FUNCTION_BLOCK "FB_GL_PROGRAM"   // FB5, GRAPH_PLUS
{ S7_Optimized_Access := 'TRUE' }
VERSION : 0.1
   VAR_INPUT
      OFF_SQ : Bool := false;   // Turn sequence off
      INIT_SQ : Bool := false;   // Set sequence to initial state
      ACK_EF : Bool := false;   // Acknowledge all errors and faults
      S_PREV : Bool := false;   // Output previous step in parameter S_NO
      S_NEXT : Bool := false;   // Indicate next step in parameter S_NO
      SW_AUTO : Bool := false;   // Automatic mode
      SW_TAP : Bool := false;   // Semiautomatic/switch with transition
      SW_TOP : Bool := false;   // Semiautomatic/ignore transition
      SW_MAN : Bool := false;   // Manual mode
      S_SEL : Int := 0;   // Select step to be output to S_NO
      S_ON : Bool := false;   // Activate step indicated in S_NO
      S_OFF : Bool := false;   // Deactivate step indicated S_NO
      T_PUSH : Bool := false;   // Enable transition to switch in semi automatic mode
   END_VAR
   VAR_OUTPUT
      S_NO : Int := 0;   // Step number
      S_MORE : Bool := false;   // More steps are available and can be shown in S_NO
      S_ACTIVE : Bool := false;   // Step indicated in S_NO is active
      ERR_FLT : Bool := false;   // Interlock or supervision group error
      AUTO_ON : Bool := false;   // Automatic mode is active
      TAP_ON : Bool := false;   // Semiautomatic mode/step with transition enabled
      TOP_ON : Bool := false;   // Semiautomatic mode/ignore transition enabled
      MAN_ON : Bool := false;   // Manual mode is active
   END_VAR
   VAR
      T_ON : Array[0..125] of TON_TIME;
   END_VAR
   VAR RETAIN
      StevecKosov : DInt;
   END_VAR
   VAR
      HMI_INFO : Array[0..34] of UInt;
      IF_PAR : G7_IfParPlus_V6;
      RT_DATA : G7_RTDataPlus_V6;   // Internal data area
      Trans9 : G7_TransitionPlus_V6;   // Transition structure
      Trans18 : G7_TransitionPlus_V6;   // Transition structure
      Trans19 : G7_TransitionPlus_V6;   // Transition structure
      Trans20 : G7_TransitionPlus_V6;   // Transition structure
      Trans22 : G7_TransitionPlus_V6;   // Transition structure
      Trans23 : G7_TransitionPlus_V6;   // Transition structure
      Trans24 : G7_TransitionPlus_V6;   // Transition structure
      Trans26 : G7_TransitionPlus_V6;   // Transition structure
      Trans28 : G7_TransitionPlus_V6;   // Transition structure
      Trans29 : G7_TransitionPlus_V6;   // Transition structure
      Trans30 : G7_TransitionPlus_V6;   // Transition structure
      Trans31 : G7_TransitionPlus_V6;   // Transition structure
      Trans32 : G7_TransitionPlus_V6;   // Transition structure
      Trans33 : G7_TransitionPlus_V6;   // Transition structure
      Trans34 : G7_TransitionPlus_V6;   // Transition structure
      Trans35 : G7_TransitionPlus_V6;   // Transition structure
      Trans36 : G7_TransitionPlus_V6;   // Transition structure
      Trans37 : G7_TransitionPlus_V6;   // Transition structure
      Trans38 : G7_TransitionPlus_V6;   // Transition structure
      Trans39 : G7_TransitionPlus_V6;   // Transition structure
      Trans40 : G7_TransitionPlus_V6;   // Transition structure
      Trans41 : G7_TransitionPlus_V6;   // Transition structure
      Trans42 : G7_TransitionPlus_V6;   // Transition structure
      Trans43 : G7_TransitionPlus_V6;   // Transition structure
      Trans44 : G7_TransitionPlus_V6;   // Transition structure
      Trans45 : G7_TransitionPlus_V6;   // Transition structure
      Trans46 : G7_TransitionPlus_V6;   // Transition structure
      Trans47 : G7_TransitionPlus_V6;   // Transition structure
      Trans48 : G7_TransitionPlus_V6;   // Transition structure
      Trans49 : G7_TransitionPlus_V6;   // Transition structure
      Trans50 : G7_TransitionPlus_V6;   // Transition structure
      Trans51 : G7_TransitionPlus_V6;   // Transition structure
      Trans52 : G7_TransitionPlus_V6;   // Transition structure
      Trans53 : G7_TransitionPlus_V6;   // Transition structure
      Trans54 : G7_TransitionPlus_V6;   // Transition structure
      Trans55 : G7_TransitionPlus_V6;   // Transition structure
      Trans56 : G7_TransitionPlus_V6;   // Transition structure
      Trans58 : G7_TransitionPlus_V6;   // Transition structure
      Trans59 : G7_TransitionPlus_V6;   // Transition structure
      Trans60 : G7_TransitionPlus_V6;   // Transition structure
      Trans61 : G7_TransitionPlus_V6;   // Transition structure
      Trans62 : G7_TransitionPlus_V6;   // Transition structure
      Trans64 : G7_TransitionPlus_V6;   // Transition structure
      Step1 : G7_StepPlus_V6;   // Step structure
      "RESET VSEGA" : G7_StepPlus_V6;   // Step structure
      "Zapiranje klešč" : G7_StepPlus_V6;   // Step structure
      "Vstavljanje v mizo" : G7_StepPlus_V6;   // Step structure
      "Odpri Držanje komada" : G7_StepPlus_V6;   // Step structure
      "Zapiranje klešč_1" : G7_StepPlus_V6;   // Step structure
      "Odpri klešče" : G7_StepPlus_V6;   // Step structure
      "DRŽI IZDELEK" : G7_StepPlus_V6;   // Step structure
      "VRAČANJE NAZAJ" : G7_StepPlus_V6;   // Step structure
      "ZAVRTI MIZO" : G7_StepPlus_V6;   // Step structure
      "ZAKLEP KONUSA" : G7_StepPlus_V6;   // Step structure
      "NALAGANJE PLOŠČICE/KOMADA" : G7_StepPlus_V6;   // Step structure
      "Odpri Držanje komada_1" : G7_StepPlus_V6;   // Step structure
      "PODAJANJE PLOŠČICE" : G7_StepPlus_V6;   // Step structure
      "Vstavljanje v mizo_1" : G7_StepPlus_V6;   // Step structure
      Step16 : G7_StepPlus_V6;   // Step structure
      "Poravnava nazaj" : G7_StepPlus_V6;   // Step structure
      "Spust Elektrode" : G7_StepPlus_V6;   // Step structure
      Varjenje : G7_StepPlus_V6;   // Step structure
      "Dvig elektrode" : G7_StepPlus_V6;   // Step structure
      "Odpri klešče_1" : G7_StepPlus_V6;   // Step structure
      "Odmik konusa" : G7_StepPlus_V6;   // Step structure
      VrtenjeVarilniELektrode : G7_StepPlus_V6;   // Step structure
      "POZ ZAVARJENO" : G7_StepPlus_V6;   // Step structure
      "IZMET KOSOV" : G7_StepPlus_V6;   // Step structure
      "Odmik vilic" : G7_StepPlus_V6;   // Step structure
      REZANJE : G7_StepPlus_V6;   // Step structure
      Step30 : G7_StepPlus_V6;   // Step structure
      "ZAČETEK NOVEGA CIKLA" : G7_StepPlus_V6;   // Step structure
      IZMET : G7_StepPlus_V6;   // Step structure
      "DRŽI IZDELEK_1" : G7_StepPlus_V6;   // Step structure
      "VRAČANJE NAZAJ_1" : G7_StepPlus_V6;   // Step structure
      "Zakasnitev varjenja" : G7_StepPlus_V6;   // Step structure
      Step36 : G7_StepPlus_V6;   // Step structure
      Step37 : G7_StepPlus_V6;   // Step structure
      Step38 : G7_StepPlus_V6;   // Step structure
      "ZAKLEP KONUSA_1" : G7_StepPlus_V6;   // Step structure
      Step40 : G7_StepPlus_V6;   // Step structure
      Step41 : G7_StepPlus_V6;   // Step structure
      Step42 : G7_StepPlus_V6;   // Step structure
      Step43 : G7_StepPlus_V6;   // Step structure
      "Izdelek ni bil prisoten" : G7_StepPlus_V6;   // Step structure
      Step45 : G7_StepPlus_V6;   // Step structure
      "Poravnava Naprej_1" : G7_StepPlus_V6;   // Step structure
      PODAJANJE_1 : G7_StepPlus_V6;   // Step structure
      "Vlaganje ploščice_1" : G7_StepPlus_V6;   // Step structure
      Step49 : G7_StepPlus_V6;   // Step structure
      "ZVAR NOK" : G7_StepPlus_V6;   // Step structure
      "Zvar  OK" : G7_StepPlus_V6;   // Step structure
      Step52 : G7_StepPlus_V6;   // Step structure
      Step53 : G7_StepPlus_V6;   // Step structure
      Step54 : G7_StepPlus_V6;   // Step structure
      SINI : Array[0..27] of USInt;
      LSTT : Array[0..42] of USInt;
      ATAJ : Array[0..42] of USInt;
      ATAB : Array[0..42] of USInt;
      PSTT : Array[0..42] of USInt;
      NSTT : Array[0..42] of USInt;
      ASSJ : Array[0..51] of USInt;
      ASSB : Array[0..51] of USInt;
      PTTS : Array[0..51] of USInt;
      NTTS : Array[0..51] of USInt;
      SW_SQTS : Array[0..51] of USInt;
      SWITCH : Array[0..171] of USInt;
      TVX : Array[0..35] of USInt;
      TTX : Array[0..35] of USInt;
      TSX : Array[0..27] of USInt;
      S00X : Array[0..27] of USInt;
      SOFFX : Array[0..27] of USInt;
      SONX : Array[0..27] of USInt;
      SAX : Array[0..27] of USInt;
      SERRX : Array[0..52] of USInt;
      SMX : Array[0..52] of USInt;
      S0X : Array[0..52] of USInt;
      S1X : Array[0..52] of USInt;
      IL_ALARM_INST : Diag_Alarm;
      SUP_ALARM_INST : Diag_Alarm;
      STEP_TIME_ALARM_INST : Diag_Alarm;
      IEC_TIMER_INST : IEC_TIMER;
      TRANSACTION_FLAG : Bool := false;
   END_VAR
   VAR_TEMP
      onemogoci : Bool;
   END_VAR
   VAR_TEMP   // added for the SCL form of the ladder/FBD networks
      _w1 : Bool;
      _w2 : Bool;
   END_VAR
   // SINI[0] := 2;
   // LSTT[0] := 255;
   // LSTT[1] := 255;
   // ATAJ[1] := 1;
   // ATAJ[2] := 2;
   // ATAB[1] := 1;
   // ATAB[2] := 2;
   // PSTT[1] := 17;
   // PSTT[2] := 32;
   // NSTT[0] := 1;
   // NSTT[1] := 16;
   // ASSJ[1] := 1;
   // ASSJ[2] := 4;
   // ASSB[1] := 1;
   // ASSB[2] := 4;
   // PTTS[0] := 255;
   // PTTS[12] := 24;
   // NTTS[1] := 8;
   // NTTS[2] := 11;
   // TVX[0] := 16#1;
   // TTX[0] := 16#1;
   // TSX[0] := 16#1;
   // S00X[0] := 16#1;
   // SOFFX[0] := 16#1;
   // SONX[0] := 16#1;
   // SAX[0] := 16#1;
   // SERRX[0] := 16#1;
   // SMX[0] := 16#1;
   // S0X[0] := 16#1;
   // S1X[0] := 16#1;
   // LSTT[3] := 255;
   // LSTT[2] := 255;
   // ATAJ[3] := 3;
   // ATAJ[4] := 4;
   // ATAB[3] := 3;
   // ATAB[4] := 4;
   // PSTT[3] := 19;
   // PSTT[4] := 27;
   // NSTT[2] := 19;
   // NSTT[3] := 22;
   // ASSJ[3] := 3;
   // ASSJ[4] := 2;
   // ASSB[3] := 3;
   // ASSB[4] := 2;
   // PTTS[3] := 11;
   // PTTS[4] := 32;
   // NTTS[3] := 12;
   // NTTS[4] := 11;
   // LSTT[4] := 255;
   // ATAJ[5] := 5;
   // ATAB[5] := 5;
   // PSTT[5] := 18;
   // NSTT[4] := 23;
   // ASSJ[5] := 12;
   // ASSB[5] := 12;
   // PTTS[5] := 24;
   // NTTS[5] := 13;
   // LSTT[6] := 255;
   // ATAJ[6] := 6;
   // ATAB[6] := 6;
   // PSTT[6] := 24;
   // NSTT[6] := 17;
   // ASSJ[6] := 7;
   // ASSB[6] := 7;
   // PTTS[6] := 12;
   // NTTS[6] := 14;
   // LSTT[5] := 255;
   // ATAJ[7] := 7;
   // ATAB[7] := 7;
   // PSTT[7] := 16;
   // NSTT[5] := 27;
   // ASSJ[7] := 6;
   // ASSB[7] := 6;
   // PTTS[7] := 12;
   // NTTS[7] := 14;
   // LSTT[7] := 255;
   // ATAJ[8] := 8;
   // ATAB[8] := 8;
   // PSTT[8] := 1;
   // NSTT[7] := 18;
   // ASSJ[8] := 21;
   // ASSB[8] := 21;
   // PTTS[8] := 14;
   // NTTS[8] := 21;
   // LSTT[8] := 255;
   // ATAJ[9] := 9;
   // ATAB[9] := 9;
   // PSTT[9] := 23;
   // NSTT[8] := 29;
   // ASSJ[9] := 33;
   // ASSB[9] := 33;
   // PTTS[9] := 21;
   // NTTS[9] := 23;
   // LSTT[9] := 255;
   // ATAJ[10] := 10;
   // ATAB[10] := 10;
   // PSTT[10] := 42;
   // NSTT[9] := 15;
   // ASSJ[10] := 43;
   // ASSJ[11] := 11;
   // ASSB[10] := 43;
   // ASSB[11] := 11;
   // PTTS[10] := 17;
   // PTTS[11] := 26;
   // NTTS[10] := 6;
   // NTTS[11] := 19;
   // LSTT[10] := 255;
   // NSTT[10] := 255;
   // SWITCH[161] := 65;
   // SINI[2] := 255;
   // SINI[3] := 255;
   // ASSB[12] := 36;
   // ASSJ[12] := 36;
   // NSTT[11] := 3;
   // PSTT[11] := 2;
   // ATAB[11] := 11;
   // ATAJ[11] := 11;
   // LSTT[11] := 255;
   // SW_SQTS[24] := 18;
   // NTTS[24] := 6;
   // LSTT[23] := 255;
   // ASSJ[24] := 10;
   // PTTS[24] := 17;
   // SINI[15] := 255;
   // SINI[14] := 255;
   // SWITCH[164] := 8;
   // SW_SQTS[4] := 3;
   // SW_SQTS[23] := 12;
   // SW_SQTS[14] := 11;
   // NTTS[12] := 13;
   // PTTS[2] := 32;
   // SW_SQTS[8] := 7;
   // SW_SQTS[9] := 8;
   // ASSB[24] := 10;
   // SWITCH[94] := 9;
   // NTTS[21] := 21;
   // PTTS[21] := 14;
   // ASSJ[21] := 8;
   // ASSB[21] := 8;
   // LSTT[12] := 255;
   // ATAJ[12] := 12;
   // ATAB[12] := 12;
   // PSTT[12] := 3;
   // NSTT[12] := 6;
   // ASSJ[13] := 13;
   // ASSB[13] := 13;
   // PTTS[13] := 19;
   // NTTS[13] := 18;
   // LSTT[13] := 255;
   // ATAJ[13] := 13;
   // ATAB[13] := 13;
   // PSTT[13] := 5;
   // NSTT[13] := 14;
   // ASSJ[14] := 14;
   // ASSB[14] := 14;
   // PTTS[14] := 13;
   // NTTS[14] := 15;
   // LSTT[14] := 255;
   // ATAJ[14] := 29;
   // ATAB[14] := 14;
   // PSTT[14] := 6;
   // NSTT[14] := 8;
   // ASSJ[15] := 15;
   // ASSB[15] := 15;
   // PTTS[15] := 9;
   // NTTS[15] := 30;
   // SINI[4] := 255;
   // SINI[5] := 255;
   // ASSJ[16] := 25;
   // ASSB[16] := 25;
   // PTTS[16] := 1;
   // NTTS[16] := 7;
   // SW_SQTS[2] := 1;
   // SW_SQTS[3] := 2;
   // SW_SQTS[5] := 4;
   // SW_SQTS[6] := 5;
   // SW_SQTS[7] := 6;
   // SW_SQTS[12] := 10;
   // SW_SQTS[21] := 17;
   // SW_SQTS[26] := 20;
   // SW_SQTS[15] := 12;
   // SW_SQTS[16] := 13;
   // SWITCH[103] := 24;
   // SINI[6] := 255;
   // SINI[7] := 255;
   // LSTT[15] := 255;
   // ATAJ[15] := 15;
   // ATAB[15] := 15;
   // PSTT[15] := 14;
   // NSTT[15] := 39;
   // ASSJ[17] := 17;
   // ASSJ[18] := 18;
   // ASSB[17] := 17;
   // ASSB[18] := 49;
   // PTTS[17] := 6;
   // PTTS[18] := 7;
   // NTTS[17] := 1;
   // NTTS[18] := 5;
   // SW_SQTS[17] := 14;
   // SW_SQTS[18] := 12;
   // LSTT[16] := 255;
   // ATAJ[16] := 16;
   // ATAB[16] := 16;
   // PSTT[16] := 44;
   // NSTT[16] := 50;
   // ASSJ[19] := 19;
   // ASSB[19] := 19;
   // PTTS[19] := 2;
   // NTTS[19] := 3;
   // SW_SQTS[19] := 15;
   // NSTT[17] := 24;
   // PSTT[17] := 34;
   // ATAJ[17] := 17;
   // LSTT[17] := 255;
   // ASSJ[20] := 30;
   // ASSB[20] := 30;
   // PTTS[20] := 34;
   // NTTS[20] := 20;
   // SW_SQTS[20] := 16;
   // SINI[8] := 255;
   // SINI[9] := 255;
   // ASSB[32] := 32;
   // ASSJ[32] := 32;
   // NTTS[27] := 4;
   // ASSJ[22] := 22;
   // ASSB[22] := 22;
   // PTTS[22] := 3;
   // NTTS[22] := 22;
   // SW_SQTS[22] := 15;
   // SWITCH[53] := 134;
   // ATAB[23] := 35;
   // LSTT[18] := 255;
   // ATAJ[18] := 18;
   // ATAB[18] := 18;
   // PSTT[18] := 13;
   // NSTT[18] := 28;
   // ASSJ[23] := 23;
   // ASSB[23] := 23;
   // PTTS[23] := 4;
   // NTTS[23] := 9;
   // SINI[22] := 255;
   // SWITCH[142] := 8;
   // SWITCH[144] := 112;
   // NSTT[19] := 13;
   // PSTT[19] := 11;
   // ATAB[19] := 19;
   // ATAJ[19] := 19;
   // LSTT[19] := 255;
   // SWITCH[123] := 4;
   // SW_SQTS[33] := 23;
   // NTTS[33] := 23;
   // PTTS[33] := 21;
   // ASSB[33] := 9;
   // SWITCH[59] := 4;
   // ASSJ[33] := 9;
   // LSTT[20] := 255;
   // LSTT[21] := 255;
   // ATAJ[20] := 33;
   // ATAJ[21] := 21;
   // ATAB[20] := 20;
   // ATAB[21] := 21;
   // PSTT[20] := 20;
   // PSTT[21] := 8;
   // NSTT[20] := 31;
   // NSTT[21] := 9;
   // ASSJ[25] := 31;
   // ASSJ[26] := 26;
   // ASSB[25] := 16;
   // ASSB[26] := 42;
   // PTTS[25] := 1;
   // PTTS[26] := 41;
   // NTTS[25] := 7;
   // NTTS[26] := 40;
   // SW_SQTS[25] := 19;
   // PSTT[23] := 9;
   // ATAJ[23] := 23;
   // LSTT[22] := 255;
   // ATAJ[22] := 22;
   // ATAB[22] := 22;
   // PSTT[22] := 22;
   // NSTT[22] := 46;
   // PTTS[27] := 5;
   // ASSB[27] := 27;
   // ASSJ[27] := 27;
   // NSTT[23] := 34;
   // SINI[18] := 255;
   // SWITCH[58] := 1;
   // SWITCH[141] := 4;
   // SINI[17] := 255;
   // PTTS[29] := 8;
   // SWITCH[85] := 132;
   // SWITCH[60] := 33;
   // SWITCH[43] := 161;
   // SWITCH[84] := 56;
   // NTTS[32] := 2;
   // SW_SQTS[32] := 15;
   // SWITCH[79] := 16;
   // PTTS[32] := 39;
   // SINI[10] := 255;
   // SINI[11] := 255;
   // SINI[12] := 255;
   // SINI[13] := 255;
   // LSTT[24] := 255;
   // LSTT[25] := 255;
   // LSTT[26] := 255;
   // ATAJ[24] := 24;
   // ATAJ[25] := 25;
   // ATAJ[26] := 26;
   // ATAB[24] := 33;
   // ATAB[25] := 27;
   // ATAB[26] := 26;
   // PSTT[24] := 37;
   // PSTT[25] := 35;
   // PSTT[26] := 29;
   // NSTT[24] := 5;
   // NSTT[25] := 40;
   // NSTT[26] := 11;
   // ASSJ[28] := 28;
   // ASSJ[29] := 29;
   // ASSJ[30] := 20;
   // ASSJ[31] := 16;
   // NSTT[28] := 35;
   // PSTT[28] := 28;
   // ASSB[28] := 28;
   // ASSB[29] := 29;
   // ASSB[30] := 20;
   // ASSB[31] := 31;
   // ATAB[28] := 28;
   // ATAJ[28] := 28;
   // PTTS[28] := 18;
   // PTTS[31] := 20;
   // PTTS[30] := 34;
   // LSTT[28] := 255;
   // NTTS[28] := 28;
   // NTTS[29] := 26;
   // NTTS[30] := 20;
   // NTTS[31] := 7;
   // SW_SQTS[10] := 9;
   // SW_SQTS[27] := 12;
   // SW_SQTS[37] := 26;
   // SW_SQTS[47] := 34;
   // SWITCH[44] := 204;
   // LSTT[27] := 255;
   // ATAJ[27] := 27;
   // ATAB[27] := 25;
   // PSTT[27] := 35;
   // NSTT[27] := 38;
   // SWITCH[147] := 24;
   // SWITCH[88] := 8;
   // SWITCH[99] := 26;
   // SWITCH[55] := 1;
   // SWITCH[102] := 128;
   // LSTT[29] := 255;
   // LSTT[30] := 255;
   // ATAJ[29] := 14;
   // ATAJ[30] := 30;
   // ATAB[29] := 29;
   // ATAB[30] := 37;
   // PSTT[29] := 38;
   // PSTT[30] := 15;
   // NSTT[29] := 8;
   // NSTT[30] := 48;
   // ASSJ[34] := 34;
   // ASSJ[35] := 35;
   // ASSB[34] := 37;
   // ASSB[35] := 35;
   // PTTS[34] := 23;
   // PTTS[35] := 28;
   // NTTS[34] := 17;
   // NTTS[35] := 25;
   // SW_SQTS[31] := 22;
   // SW_SQTS[34] := 24;
   // SW_SQTS[38] := 27;
   // NTTS[38] := 29;
   // PTTS[38] := 27;
   // ASSB[38] := 38;
   // ASSJ[38] := 38;
   // ASSJ[36] := 5;
   // ASSB[36] := 5;
   // PTTS[36] := 24;
   // NTTS[36] := 13;
   // SW_SQTS[48] := 35;
   // ASSJ[37] := 37;
   // SINI[16] := 255;
   // SWITCH[146] := 51;
   // SWITCH[105] := 224;
   // SWITCH[121] := 136;
   // SWITCH[73] := 130;
   // ASSB[37] := 34;
   // PTTS[37] := 23;
   // NTTS[37] := 24;
   // SW_SQTS[39] := 11;
   // SWITCH[62] := 210;
   // SWITCH[34] := 16;
   // SWITCH[91] := 3;
   // LSTT[31] := 255;
   // ATAJ[31] := 35;
   // ATAB[31] := 31;
   // PSTT[31] := 46;
   // NSTT[31] := 41;
   // ASSJ[39] := 39;
   // ASSB[39] := 39;
   // PTTS[39] := 15;
   // NTTS[39] := 34;
   // LSTT[33] := 255;
   // LSTT[32] := 255;
   // ATAJ[32] := 32;
   // ATAJ[33] := 20;
   // ATAB[32] := 32;
   // ATAB[33] := 24;
   // PSTT[32] := 40;
   // PSTT[33] := 37;
   // NSTT[32] := 2;
   // NSTT[33] := 31;
   // ASSJ[40] := 40;
   // ASSJ[41] := 41;
   // ASSB[40] := 40;
   // ASSB[41] := 41;
   // PTTS[40] := 25;
   // PTTS[41] := 31;
   // NTTS[40] := 32;
   // NTTS[41] := 36;
   // SW_SQTS[40] := 28;
   // SW_SQTS[41] := 29;
   // SWITCH[107] := 8;
   // SWITCH[152] := 2;
   // LSTT[34] := 255;
   // ATAJ[34] := 34;
   // ATAB[34] := 34;
   // PSTT[34] := 39;
   // NSTT[34] := 20;
   // LSTT[35] := 255;
   // ATAJ[35] := 31;
   // ATAB[35] := 23;
   // PSTT[35] := 9;
   // NSTT[35] := 41;
   // ASSJ[42] := 42;
   // ASSB[42] := 26;
   // PTTS[42] := 41;
   // NTTS[42] := 10;
   // SW_SQTS[42] := 30;
   // LSTT[36] := 28;
   // ATAJ[36] := 36;
   // ATAB[36] := 36;
   // PSTT[36] := 41;
   // NSTT[36] := 28;
   // SWITCH[156] := 48;
   // ASSJ[43] := 45;
   // ASSB[43] := 45;
   // PTTS[43] := 17;
   // NTTS[43] := 6;
   // SW_SQTS[43] := 31;
   // SWITCH[87] := 14;
   // SWITCH[96] := 198;
   // SWITCH[138] := 32;
   // SWITCH[42] := 130;
   // SWITCH[148] := 16;
   // SWITCH[101] := 7;
   // SWITCH[71] := 128;
   // SWITCH[90] := 48;
   // SWITCH[113] := 97;
   // SWITCH[50] := 14;
   // SWITCH[46] := 64;
   // SWITCH[14] := 1;
   // ASSJ[44] := 44;
   // ASSB[44] := 24;
   // PTTS[44] := 17;
   // NTTS[44] := 16;
   // SW_SQTS[44] := 32;
   // SWITCH[66] := 67;
   // SWITCH[48] := 49;
   // SWITCH[54] := 192;
   // SWITCH[75] := 98;
   // SWITCH[63] := 12;
   // SWITCH[116] := 194;
   // LSTT[37] := 255;
   // LSTT[38] := 255;
   // LSTT[39] := 255;
   // ATAJ[37] := 37;
   // ATAJ[38] := 39;
   // ATAJ[39] := 38;
   // ATAB[37] := 30;
   // ATAB[38] := 38;
   // ATAB[39] := 39;
   // PSTT[37] := 15;
   // PSTT[38] := 47;
   // PSTT[39] := 48;
   // NSTT[37] := 47;
   // NSTT[38] := 32;
   // NSTT[39] := 32;
   // ASSJ[45] := 50;
   // ASSJ[46] := 46;
   // ASSB[45] := 44;
   // ASSB[46] := 46;
   // PTTS[45] := 17;
   // PTTS[46] := 22;
   // NTTS[45] := 6;
   // NTTS[46] := 31;
   // SW_SQTS[45] := 33;
   // SW_SQTS[46] := 15;
   // SWITCH[145] := 40;
   // SWITCH[61] := 24;
   // SWITCH[28] := 8;
   // NTTS[47] := 38;
   // PTTS[47] := 37;
   // ASSB[47] := 47;
   // SW_SQTS[30] := 21;
   // ASSJ[47] := 47;
   // LSTT[40] := 255;
   // SWITCH[117] := 140;
   // SWITCH[39] := 128;
   // ATAJ[40] := 40;
   // SWITCH[118] := 33;
   // ATAB[40] := 40;
   // SWITCH[143] := 131;
   // SWITCH[104] := 67;
   // PSTT[40] := 26;
   // SWITCH[122] := 49;
   // SWITCH[86] := 25;
   // NSTT[40] := 51;
   // SWITCH[98] := 196;
   // SWITCH[137] := 128;
   // SWITCH[89] := 150;
   // SWITCH[49] := 12;
   // SINI[20] := 255;
   // SINI[19] := 255;
   // SINI[21] := 255;
   // SINI[23] := 255;
   // SINI[24] := 255;
   // ASSJ[48] := 48;
   // ASSB[48] := 48;
   // PTTS[48] := 30;
   // NTTS[48] := 39;
   // SW_SQTS[36] := 25;
   // SWITCH[65] := 4;
   // SWITCH[140] := 36;
   // SWITCH[150] := 101;
   // SWITCH[149] := 14;
   // SWITCH[119] := 112;
   // SINI[25] := 255;
   // LSTT[41] := 255;
   // ATAJ[41] := 41;
   // ATAB[41] := 41;
   // PSTT[41] := 49;
   // NSTT[41] := 26;
   // ASSJ[49] := 49;
   // ASSB[49] := 18;
   // PTTS[49] := 7;
   // NTTS[49] := 41;
   // SW_SQTS[49] := 36;
   // SWITCH[52] := 49;
   // SWITCH[77] := 129;
   // SWITCH[67] := 152;
   // SWITCH[78] := 3;
   // SWITCH[100] := 2;
   // SWITCH[114] := 6;
   // SWITCH[47] := 136;
   // SWITCH[45] := 112;
   // SWITCH[155] := 204;
   // SINI[26] := 255;
   // SWITCH[124] := 14;
   // SWITCH[151] := 134;
   // ATAB[17] := 17;
   // SWITCH[23] := 128;
   // SWITCH[22] := 56;
   // SWITCH[21] := 48;
   // SWITCH[20] := 198;
   // SWITCH[5] := 1;
   // SINI[27] := 255;
   // ASSJ[50] := 24;
   // ASSB[50] := 50;
   // PTTS[50] := 16;
   // NTTS[50] := 6;
   // SW_SQTS[50] := 32;
   // SWITCH[68] := 1;
   // SWITCH[153] := 194;
   // SWITCH[154] := 161;
   // SWITCH[159] := 64;
   // SWITCH[165] := 32;
   // SWITCH[166] := 8;
   // SWITCH[168] := 9;
   // SWITCH[170] := 194;
   // LSTT[42] := 255;
   // ATAJ[42] := 42;
   // ATAB[42] := 42;
   // PSTT[42] := 51;
   // NSTT[42] := 255;
   // ASSJ[51] := 51;
   // ASSB[51] := 51;
   // PTTS[51] := 40;
   // NTTS[51] := 42;
   // SW_SQTS[51] := 20;
   // SWITCH[76] := 44;
   // SWITCH[83] := 64;
   // SWITCH[112] := 12;
   // SWITCH[111] := 16;
   // SWITCH[136] := 32;
   // SWITCH[19] := 96;
BEGIN
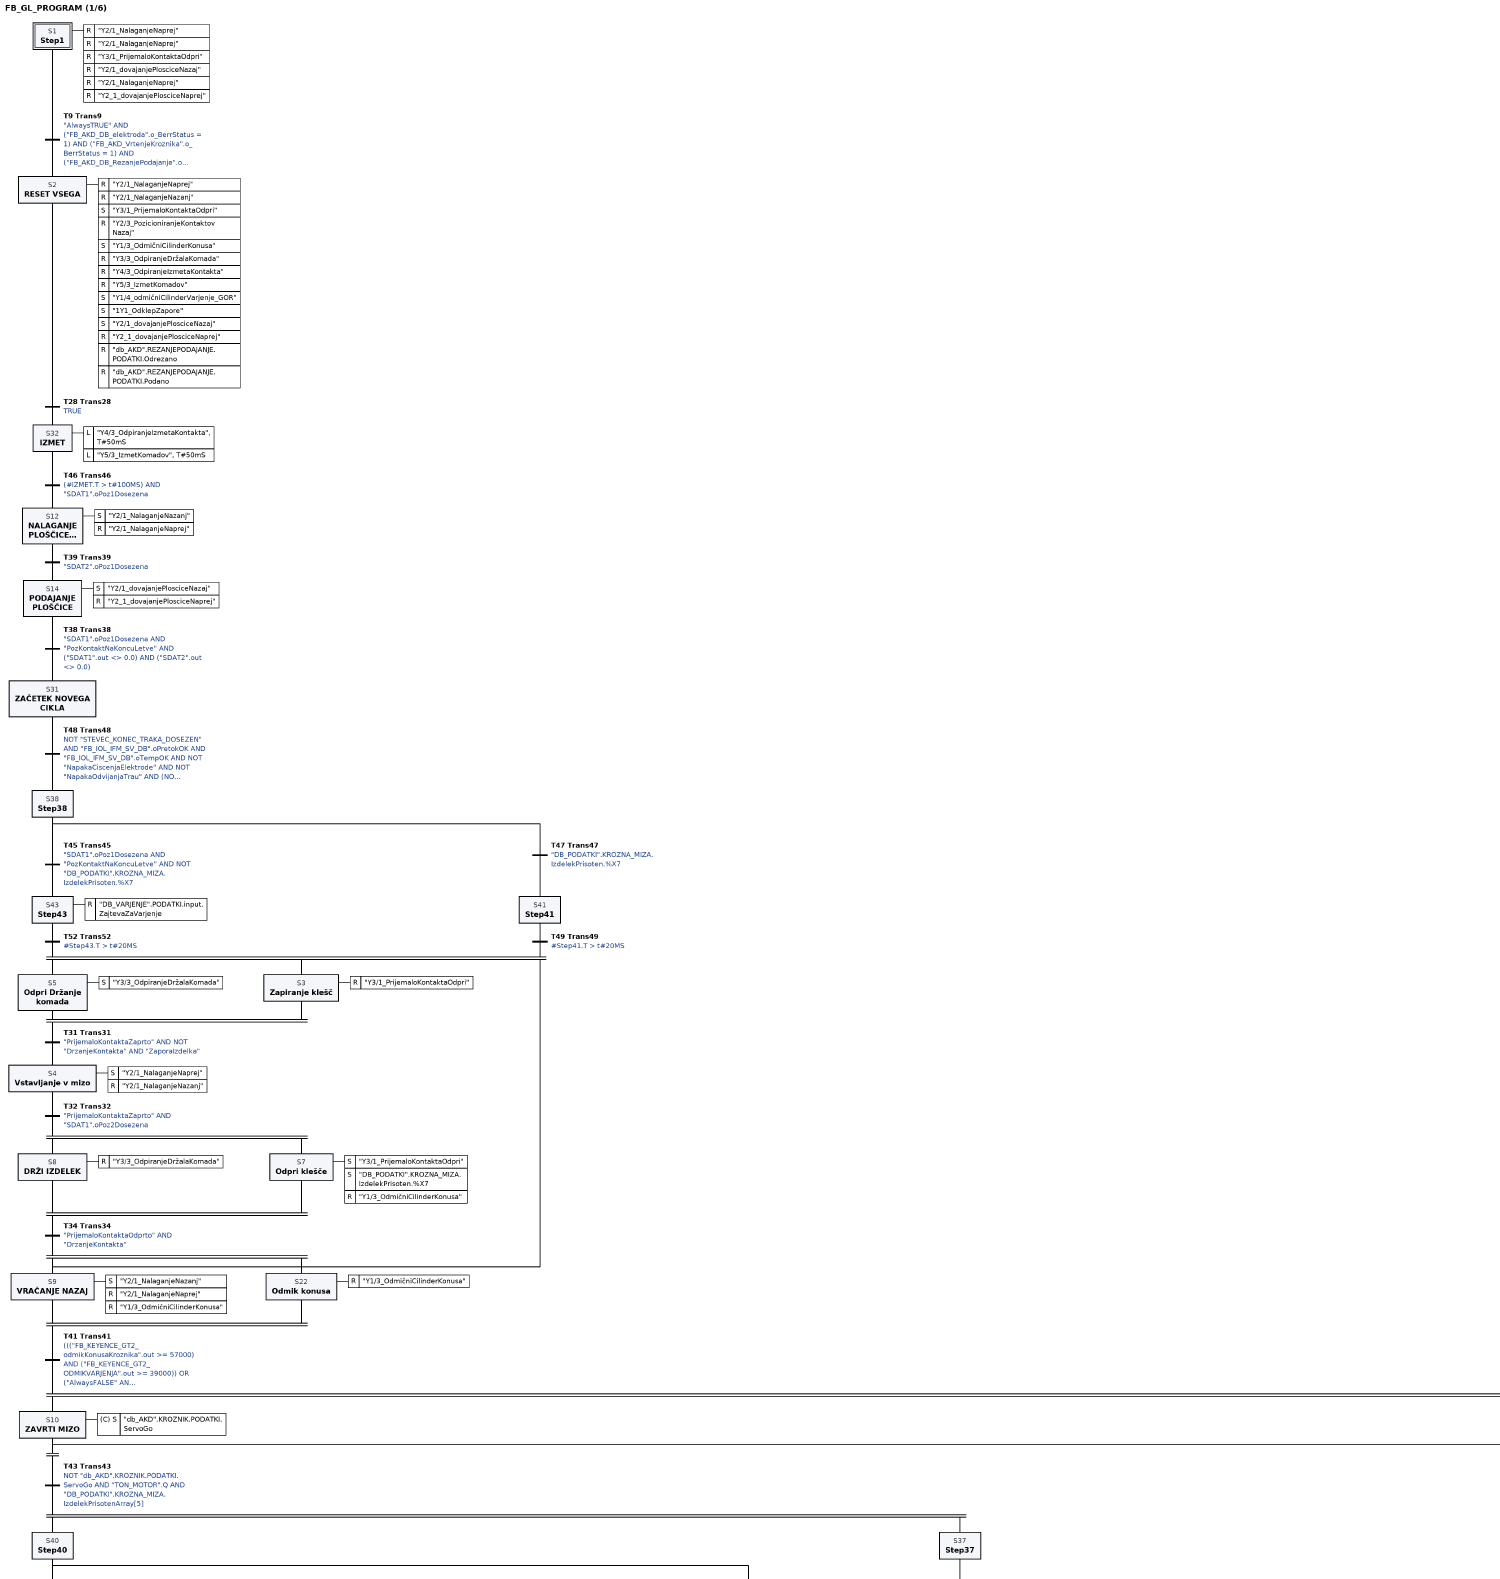
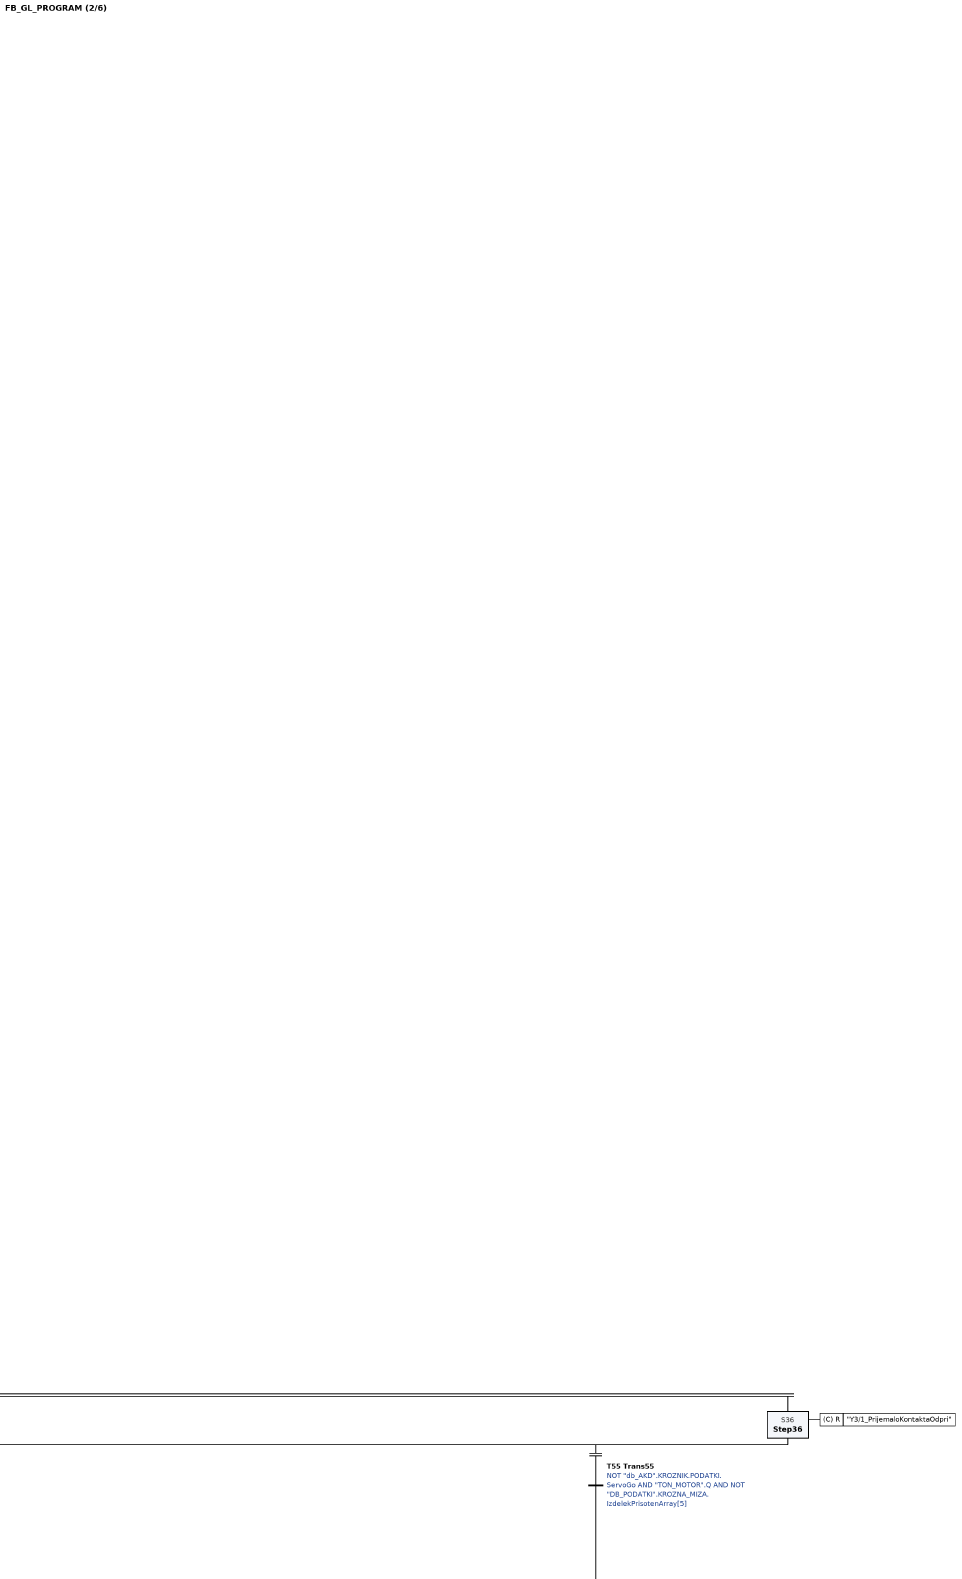
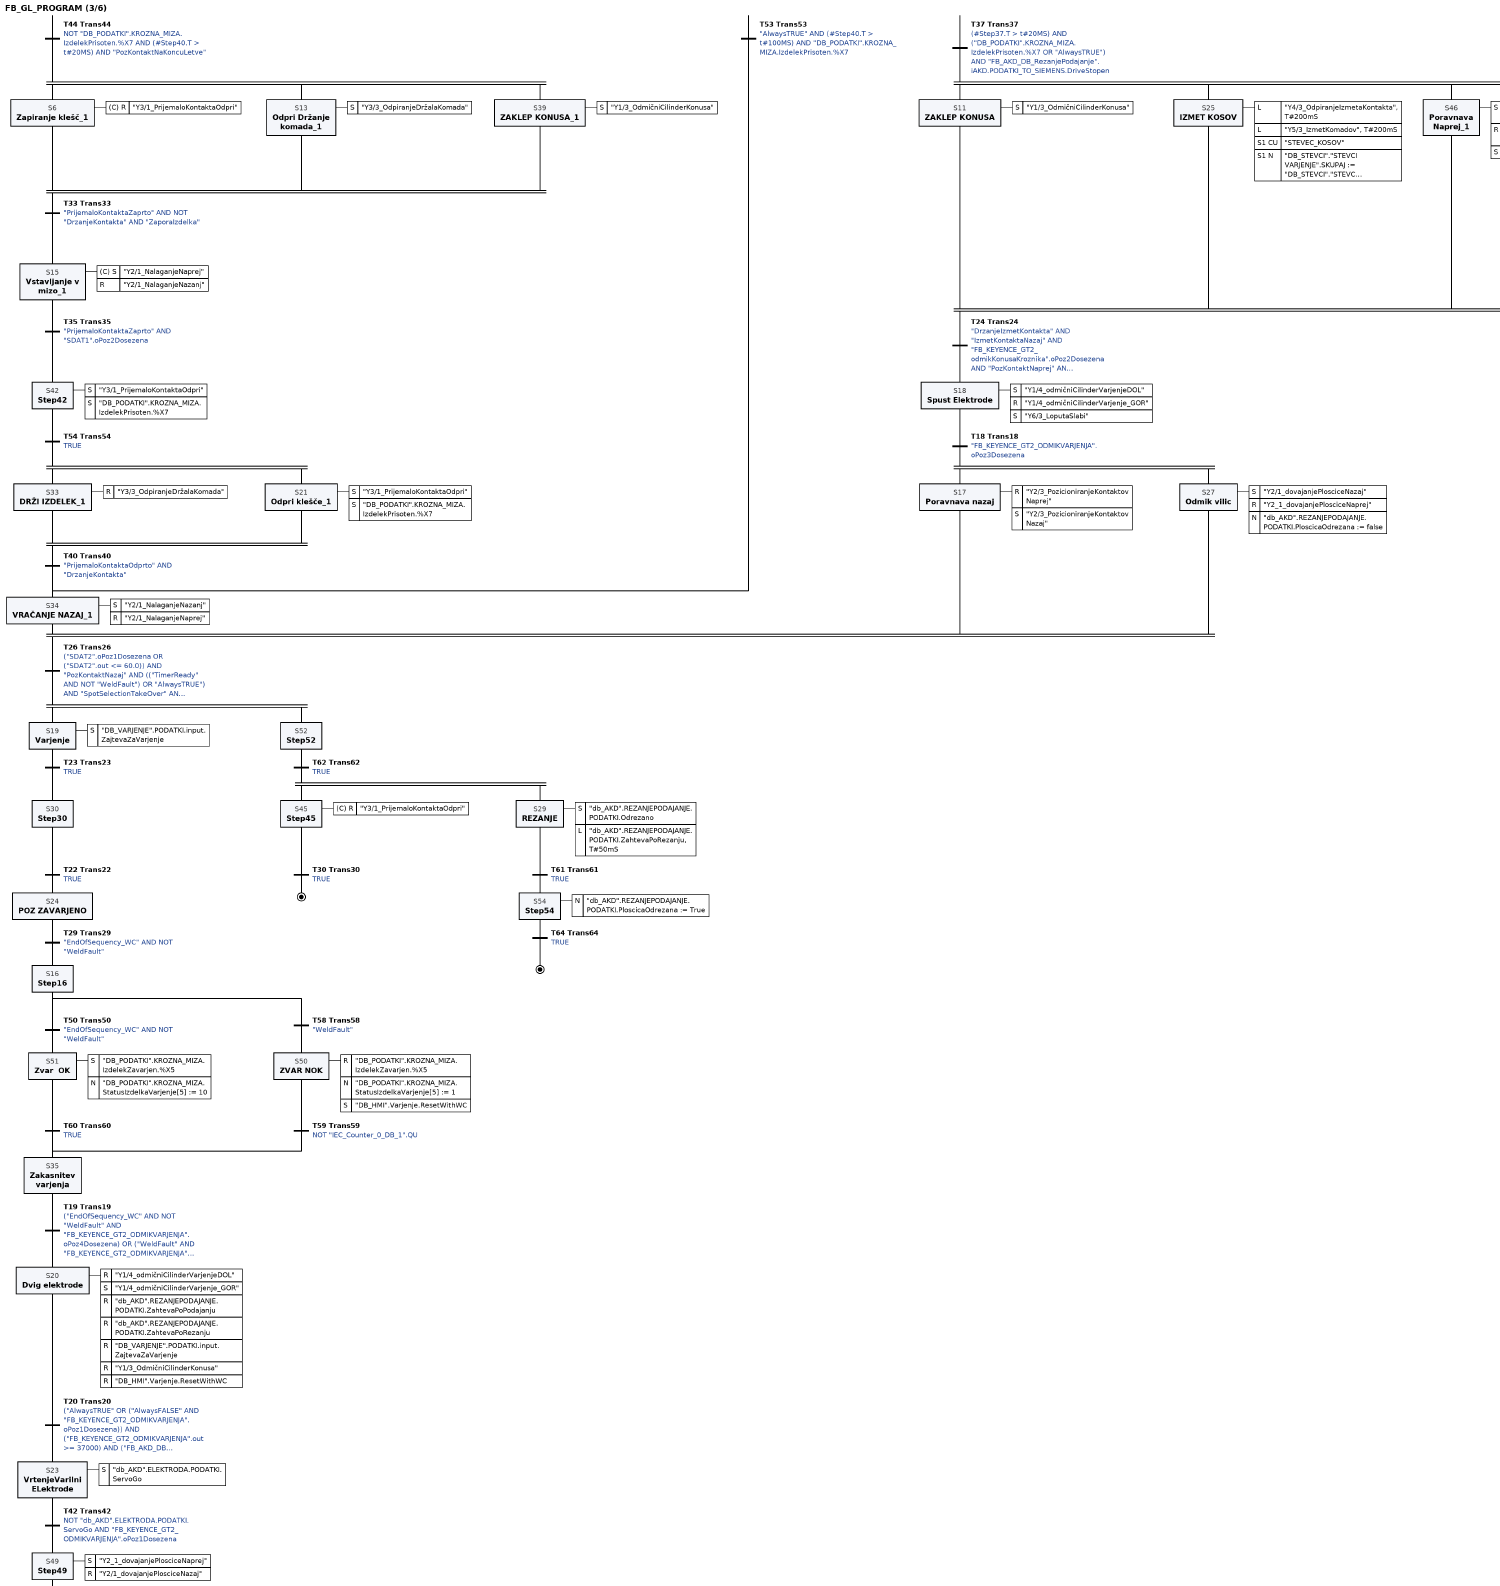
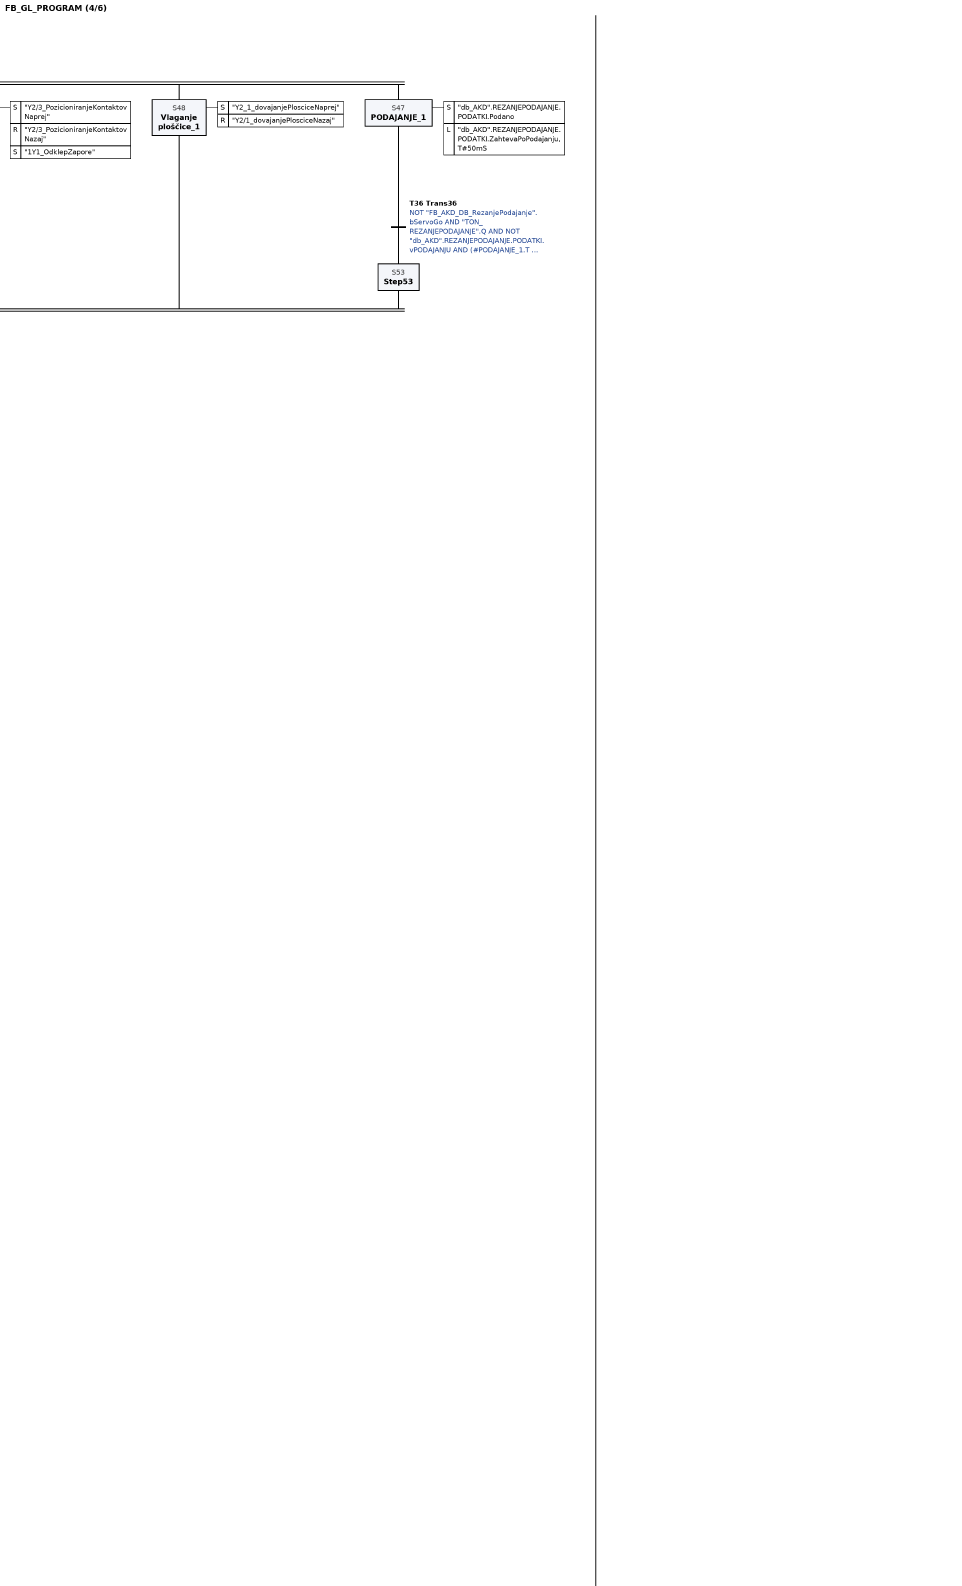
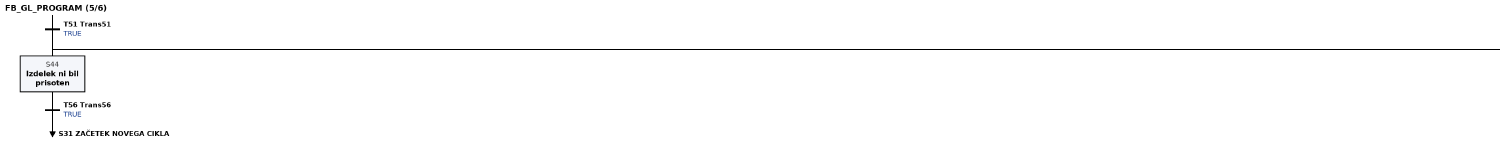
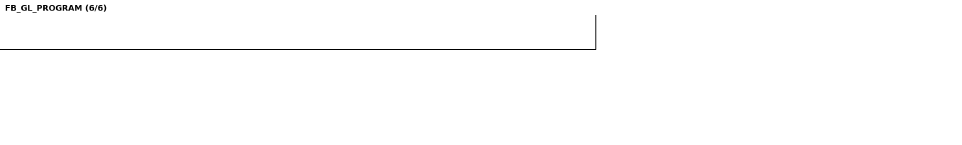
   // permanent pre-instructions
   NETWORK 1
      "TON_MOTOR".TON(IN := NOT "db_AKD".KROZNIK.PODATKI.ServoGo, PT := T#20mS);
   NETWORK 2
      "TON_REZANJEPODAJANJE".TON(IN := NOT "db_AKD".REZANJEPODAJANJE.PODATKI.ServoGO, PT := T#20mS);
   NETWORK 3
   TITLE = Generiranje Napak
      "FB_Alarms_DB".I_Alarm_1 := ("SDAT1".out = 0.0) OR ("SDAT2".out = 0.0);
   NETWORK 4
      "IEC_Counter_0_DB_1".CTU(CU := #"ZVAR NOK".X,
                              R := ("IEC_Counter_0_DB_1".QU AND "ResetNapake") OR (NOT "IEC_Counter_0_DB_1".QU AND #"Zakasnitev varjenja".X),
                              PV := 2);
   NETWORK 5
      "Y6/3_LoputaDobri" := "DB_PODATKI".KROZNA_MIZA.IzdelekPrisotenArray[1] AND "DB_PODATKI".KROZNA_MIZA.IzdelekKameraOk.%X1 AND ("DB_PODATKI".KROZNA_MIZA.StatusIzdelkaVarjenje[1] = 10) AND "AlwaysFALSE";
      "Y6/3_LoputaSlabi" := NOT "Y6/3_LoputaDobri";

   // sequencer 1
   INITIAL_STEP Step1:   // S1, max time T#10S, warning time T#7S
      supervision V := (("FB_AKD_DB_elektroda".o_BerrStatus <> 1) OR ("FB_AKD_VrtenjeKroznika".o_BerrStatus <> 1) OR ("FB_AKD_DB_RezanjePodajanje".o_BerrStatus <> 1)) AND (#Step1.T > t#2000MS);
              R    "Y2/1_NalaganjeNaprej"
              R    "Y2/1_NalaganjeNaprej"
              R    "Y3/1_PrijemaloKontaktaOdpri"
              R    "Y2/1_dovajanjePlosciceNazaj"
              R    "Y2/1_NalaganjeNaprej"
              R    "Y2_1_dovajanjePlosciceNaprej"
   END_STEP
   TRANSITION Trans9 FROM Step1 TO "RESET VSEGA"   // T9
      := "AlwaysTRUE" AND ("FB_AKD_DB_elektroda".o_BerrStatus = 1) AND ("FB_AKD_VrtenjeKroznika".o_BerrStatus = 1) AND ("FB_AKD_DB_RezanjePodajanje".o_BerrStatus = 1);
   END_TRANSITION
   STEP VrtenjeVarilniELektrode:   // S23, max time T#10S, warning time T#7S
      supervision V := "db_AKD".ELEKTRODA.PODATKI.ServoGo AND (#VrtenjeVarilniELektrode.T > t#2000MS);
              S    "db_AKD".ELEKTRODA.PODATKI.ServoGo
   END_STEP
   TRANSITION Trans42 FROM VrtenjeVarilniELektrode TO Step49   // T42
      := NOT "db_AKD".ELEKTRODA.PODATKI.ServoGo AND "FB_KEYENCE_GT2_ODMIKVARJENJA".oPoz1Dosezena;
   END_TRANSITION
   STEP "POZ ZAVARJENO":   // S24, max time T#10S, warning time T#7S
      supervision V := NOT "EndOfSequency_WC" AND (#"POZ ZAVARJENO".T > t#2000MS);
   END_STEP
   TRANSITION Trans29 FROM "POZ ZAVARJENO" TO Step16   // T29
      := "EndOfSequency_WC" AND NOT "WeldFault";
   END_TRANSITION
   STEP "Spust Elektrode":   // S18, max time T#10S, warning time T#7S
      interlock C := "SDAT2".oPoz2Dosezena;
      // Spustimo elektrodo || Restiraj - ploščica ni narejena!
              S    "Y1/4_odmičniCilinderVarjenjeDOL"
              R    "Y1/4_odmičniCilinderVarjenje_GOR"
              S    "Y6/3_LoputaSlabi"
   END_STEP
   TRANSITION Trans18 FROM "Spust Elektrode" TO ("Poravnava nazaj", "Odmik vilic")   // T18: Elektroda V poziciji za varjenje
      := "FB_KEYENCE_GT2_ODMIKVARJENJA".oPoz3Dosezena;
   END_TRANSITION
   STEP Varjenje:   // S19, max time T#10S, warning time T#7S
      supervision V := (NOT "SDAT2".oPoz1Dosezena OR NOT "FB_KEYENCE_GT2_ODMIKVARJENJA".oPoz3Dosezena OR NOT "SDAT1".oPoz1Dosezena) AND (#Varjenje.T > t#2000MS);
              S    "DB_VARJENJE".PODATKI.input.ZajtevaZaVarjenje
   END_STEP
   TRANSITION Trans23 FROM Varjenje TO Step30   // T23
      := TRUE;
   END_TRANSITION
   STEP "Dvig elektrode":   // S20, max time T#10S, warning time T#7S
      supervision V := NOT "FB_KEYENCE_GT2_ODMIKVARJENJA".oPoz1Dosezena AND (#"Dvig elektrode".T > t#2000MS);
              R    "Y1/4_odmičniCilinderVarjenjeDOL"
              S    "Y1/4_odmičniCilinderVarjenje_GOR"
              R    "db_AKD".REZANJEPODAJANJE.PODATKI.ZahtevaPoPodajanju
              R    "db_AKD".REZANJEPODAJANJE.PODATKI.ZahtevaPoRezanju
              R    "DB_VARJENJE".PODATKI.input.ZajtevaZaVarjenje
              R    "Y1/3_OdmičniCilinderKonusa"
              R    "DB_HMI".Varjenje.ResetWithWC
   END_STEP
   TRANSITION Trans20 FROM "Dvig elektrode" TO VrtenjeVarilniELektrode   // T20
      := ("AlwaysTRUE" OR ("AlwaysFALSE" AND "FB_KEYENCE_GT2_ODMIKVARJENJA".oPoz1Dosezena)) AND ("FB_KEYENCE_GT2_ODMIKVARJENJA".out >= 37000) AND ("FB_AKD_DB_elektroda".o_BerrStatus = 1);
   END_TRANSITION
   STEP "IZMET KOSOV":   // S25, max time T#10S, warning time T#7S
              L    "Y4/3_OdpiranjeIzmetaKontakta",T#200mS
              L    "Y5/3_IzmetKomadov", T#200mS
          S1  CU   "STEVEC_KOSOV"
          S1  N    "DB_STEVCI"."STEVCI VARJENJE".SKUPAJ := "DB_STEVCI"."STEVCI VARJENJE".SKUPAJ + 1
   END_STEP
   STEP "Poravnava nazaj":   // S17, max time T#10S, warning time T#7S
              R    "Y2/3_PozicioniranjeKontaktovNaprej"
              S    "Y2/3_PozicioniranjeKontaktovNazaj"
   END_STEP
   STEP Step45:   // S45, max time T#10S, warning time T#7S
      interlock C := "PozKontaktNaKoncuLetve" AND "SDAT1".oPoz1Dosezena;
      supervision V := (NOT "PozKontaktNaKoncuLetve" OR NOT "SDAT1".oPoz1Dosezena) AND (#Step45.T > t#2000MS);
      (C)     R    "Y3/1_PrijemaloKontaktaOdpri"
   END_STEP
   TRANSITION Trans30 FROM Step45 TO END   // T30
      := TRUE;
   END_TRANSITION
   STEP REZANJE:   // S29, max time T#10S, warning time T#7S
              S    "db_AKD".REZANJEPODAJANJE.PODATKI.Odrezano
              L    "db_AKD".REZANJEPODAJANJE.PODATKI.ZahtevaPoRezanju,T#50mS
   END_STEP
   TRANSITION Trans61 FROM REZANJE TO Step54   // T61
      := TRUE;
   END_TRANSITION
   STEP "NALAGANJE PLOŠČICE/KOMADA":   // S12, max time T#10S, warning time T#7S
      supervision V := (NOT "SDAT2".oPoz1Dosezena OR NOT "SDAT1".oPoz1Dosezena) AND (#"NALAGANJE PLOŠČICE/KOMADA".T > t#2000MS);
      // Klešče Se ne zaletijo
              S    "Y2/1_NalaganjeNazanj"
              R    "Y2/1_NalaganjeNaprej"
   END_STEP
   TRANSITION Trans39 FROM "NALAGANJE PLOŠČICE/KOMADA" TO "PODAJANJE PLOŠČICE"   // T39
      := "SDAT2".oPoz1Dosezena;
   END_TRANSITION
   STEP "Zapiranje klešč":   // S3, max time T#10S, warning time T#7S
      supervision V := NOT "PrijemaloKontaktaZaprto" AND (#"Zapiranje klešč".T > t#2000MS);
              R    "Y3/1_PrijemaloKontaktaOdpri"
   END_STEP
   STEP "Vstavljanje v mizo":   // S4, max time T#10S, warning time T#7S
      supervision V := NOT "PrijemaloKontaktaZaprto" AND NOT "SDAT1".oPoz2Dosezena AND (#"Vstavljanje v mizo".T > t#2000MS);
              S    "Y2/1_NalaganjeNaprej"
              R    "Y2/1_NalaganjeNazanj"
   END_STEP
   TRANSITION Trans32 FROM "Vstavljanje v mizo" TO ("DRŽI IZDELEK", "Odpri klešče")   // T32
      := "PrijemaloKontaktaZaprto" AND "SDAT1".oPoz2Dosezena;
   END_TRANSITION
   STEP "Odpri Držanje komada":   // S5, max time T#10S, warning time T#7S
      supervision V := "DrzanjeKontakta" AND (#"Odpri Držanje komada".T > t#2000MS);
      // OdpriDržanjeKomada -
              S    "Y3/3_OdpiranjeDržalaKomada"
   END_STEP
   TRANSITION Trans31 FROM ("Zapiranje klešč", "Odpri Držanje komada") TO "Vstavljanje v mizo"   // T31
      := "PrijemaloKontaktaZaprto" AND NOT "DrzanjeKontakta" AND "ZaporaIzdelka";
   END_TRANSITION
   STEP "Odpri klešče":   // S7, max time T#10S, warning time T#7S
      supervision V := NOT "PrijemaloKontaktaOdprto" AND (#"Odpri klešče".T > t#2000MS);
              S    "Y3/1_PrijemaloKontaktaOdpri"
              S    "DB_PODATKI".KROZNA_MIZA.IzdelekPrisoten.%X7
              R    "Y1/3_OdmičniCilinderKonusa"
   END_STEP
   STEP "DRŽI IZDELEK":   // S8, max time T#10S, warning time T#7S
      supervision V := NOT "DrzanjeKontakta" AND (#"DRŽI IZDELEK".T > t#2000MS);